REGION Network 249: CARRIER DRIVE INTERNAL COMM ERROR
   RUNG wire#powerrail
      { S7_Templates := "SrcType := Word" } EQ_Contact(in1 := "DB101_DB_SDC_FAULTS".Carrier_Fault[37], in2 := 151)
      Coil( "DB302_HMI_Faults".Carrier37_Faults_1.%X3 )
   END_RUNG
   // the same network as SCL:
   "DB302_HMI_Faults".Carrier37_Faults_1.%X3 := "DB101_DB_SDC_FAULTS".Carrier_Fault[37] = 151;
END_REGION

REGION Network 250: CARRIER DRIVE MOTOR OVERTEMP
   RUNG wire#powerrail
      { S7_Templates := "SrcType := Word" } EQ_Contact(in1 := "DB101_DB_SDC_FAULTS".Carrier_Fault[37], in2 := 160)
      Coil( "DB302_HMI_Faults".Carrier37_Faults_1.%X4 )
   END_RUNG
   // the same network as SCL:
   "DB302_HMI_Faults".Carrier37_Faults_1.%X4 := "DB101_DB_SDC_FAULTS".Carrier_Fault[37] = 160;
END_REGION

REGION Network 251: CARRIER DRIVE MOTOR OVERCURRENT
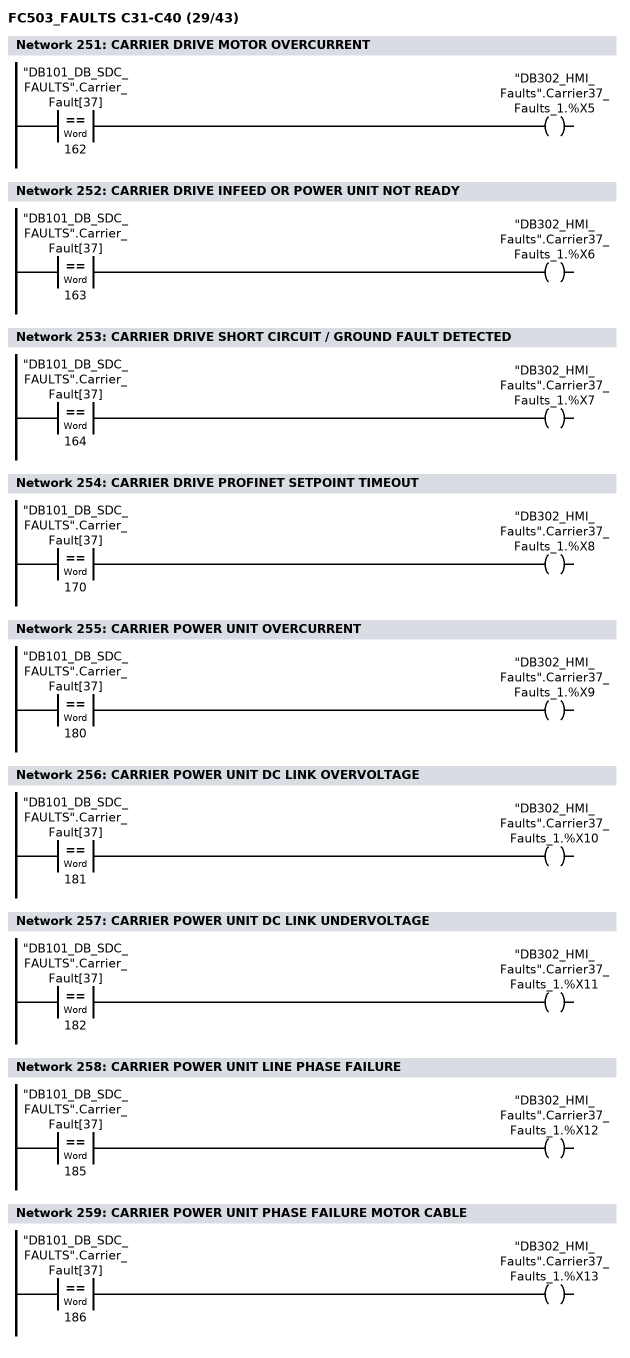
   RUNG wire#powerrail
      { S7_Templates := "SrcType := Word" } EQ_Contact(in1 := "DB101_DB_SDC_FAULTS".Carrier_Fault[37], in2 := 162)
      Coil( "DB302_HMI_Faults".Carrier37_Faults_1.%X5 )
   END_RUNG
   // the same network as SCL:
   "DB302_HMI_Faults".Carrier37_Faults_1.%X5 := "DB101_DB_SDC_FAULTS".Carrier_Fault[37] = 162;
END_REGION

REGION Network 252: CARRIER DRIVE INFEED OR POWER UNIT NOT READY
   RUNG wire#powerrail
      { S7_Templates := "SrcType := Word" } EQ_Contact(in1 := "DB101_DB_SDC_FAULTS".Carrier_Fault[37], in2 := 163)
      Coil( "DB302_HMI_Faults".Carrier37_Faults_1.%X6 )
   END_RUNG
   // the same network as SCL:
   "DB302_HMI_Faults".Carrier37_Faults_1.%X6 := "DB101_DB_SDC_FAULTS".Carrier_Fault[37] = 163;
END_REGION

REGION Network 253: CARRIER DRIVE SHORT CIRCUIT / GROUND FAULT DETECTED
   RUNG wire#powerrail
      { S7_Templates := "SrcType := Word" } EQ_Contact(in1 := "DB101_DB_SDC_FAULTS".Carrier_Fault[37], in2 := 164)
      Coil( "DB302_HMI_Faults".Carrier37_Faults_1.%X7 )
   END_RUNG
   // the same network as SCL:
   "DB302_HMI_Faults".Carrier37_Faults_1.%X7 := "DB101_DB_SDC_FAULTS".Carrier_Fault[37] = 164;
END_REGION

REGION Network 254: CARRIER DRIVE PROFINET SETPOINT TIMEOUT
   RUNG wire#powerrail
      { S7_Templates := "SrcType := Word" } EQ_Contact(in1 := "DB101_DB_SDC_FAULTS".Carrier_Fault[37], in2 := 170)
      Coil( "DB302_HMI_Faults".Carrier37_Faults_1.%X8 )
   END_RUNG
   // the same network as SCL:
   "DB302_HMI_Faults".Carrier37_Faults_1.%X8 := "DB101_DB_SDC_FAULTS".Carrier_Fault[37] = 170;
END_REGION

REGION Network 255: CARRIER POWER UNIT OVERCURRENT
   RUNG wire#powerrail
      { S7_Templates := "SrcType := Word" } EQ_Contact(in1 := "DB101_DB_SDC_FAULTS".Carrier_Fault[37], in2 := 180)
      Coil( "DB302_HMI_Faults".Carrier37_Faults_1.%X9 )
   END_RUNG
   // the same network as SCL:
   "DB302_HMI_Faults".Carrier37_Faults_1.%X9 := "DB101_DB_SDC_FAULTS".Carrier_Fault[37] = 180;
END_REGION

REGION Network 256: CARRIER POWER UNIT DC LINK OVERVOLTAGE
   RUNG wire#powerrail
      { S7_Templates := "SrcType := Word" } EQ_Contact(in1 := "DB101_DB_SDC_FAULTS".Carrier_Fault[37], in2 := 181)
      Coil( "DB302_HMI_Faults".Carrier37_Faults_1.%X10 )
   END_RUNG
   // the same network as SCL:
   "DB302_HMI_Faults".Carrier37_Faults_1.%X10 := "DB101_DB_SDC_FAULTS".Carrier_Fault[37] = 181;
END_REGION

REGION Network 257: CARRIER POWER UNIT DC LINK UNDERVOLTAGE
   RUNG wire#powerrail
      { S7_Templates := "SrcType := Word" } EQ_Contact(in1 := "DB101_DB_SDC_FAULTS".Carrier_Fault[37], in2 := 182)
      Coil( "DB302_HMI_Faults".Carrier37_Faults_1.%X11 )
   END_RUNG
   // the same network as SCL:
   "DB302_HMI_Faults".Carrier37_Faults_1.%X11 := "DB101_DB_SDC_FAULTS".Carrier_Fault[37] = 182;
END_REGION

REGION Network 258: CARRIER POWER UNIT LINE PHASE FAILURE
   RUNG wire#powerrail
      { S7_Templates := "SrcType := Word" } EQ_Contact(in1 := "DB101_DB_SDC_FAULTS".Carrier_Fault[37], in2 := 185)
      Coil( "DB302_HMI_Faults".Carrier37_Faults_1.%X12 )
   END_RUNG
   // the same network as SCL:
   "DB302_HMI_Faults".Carrier37_Faults_1.%X12 := "DB101_DB_SDC_FAULTS".Carrier_Fault[37] = 185;
END_REGION

REGION Network 259: CARRIER POWER UNIT PHASE FAILURE MOTOR CABLE
   RUNG wire#powerrail
      { S7_Templates := "SrcType := Word" } EQ_Contact(in1 := "DB101_DB_SDC_FAULTS".Carrier_Fault[37], in2 := 186)
      Coil( "DB302_HMI_Faults".Carrier37_Faults_1.%X13 )
   END_RUNG
   // the same network as SCL:
   "DB302_HMI_Faults".Carrier37_Faults_1.%X13 := "DB101_DB_SDC_FAULTS".Carrier_Fault[37] = 186;
END_REGION

REGION Network 260: CARRIER POWER UNIT GROUND FAULT
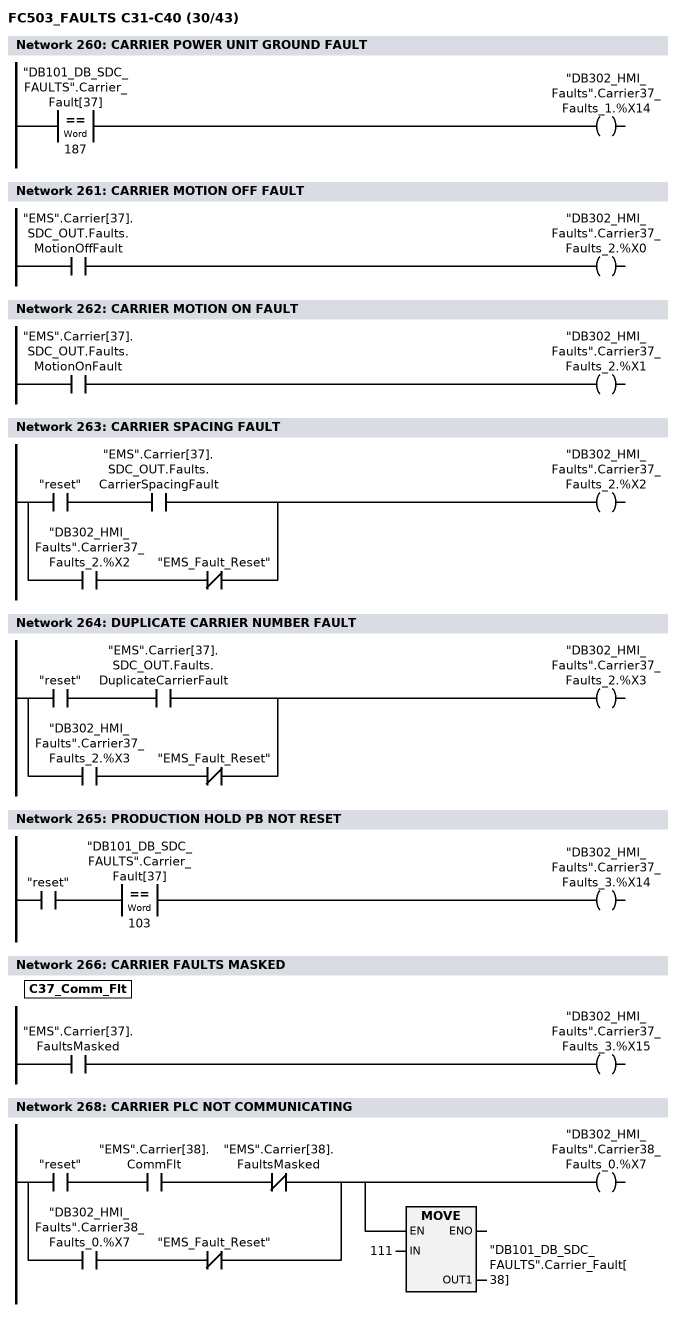
   RUNG wire#powerrail
      { S7_Templates := "SrcType := Word" } EQ_Contact(in1 := "DB101_DB_SDC_FAULTS".Carrier_Fault[37], in2 := 187)
      Coil( "DB302_HMI_Faults".Carrier37_Faults_1.%X14 )
   END_RUNG
   // the same network as SCL:
   "DB302_HMI_Faults".Carrier37_Faults_1.%X14 := "DB101_DB_SDC_FAULTS".Carrier_Fault[37] = 187;
END_REGION

REGION Network 261: CARRIER MOTION OFF FAULT
   RUNG wire#powerrail
      Contact( "EMS".Carrier[37].SDC_OUT.Faults.MotionOffFault )
      Coil( "DB302_HMI_Faults".Carrier37_Faults_2.%X0 )
   END_RUNG
   // the same network as SCL:
   "DB302_HMI_Faults".Carrier37_Faults_2.%X0 := "EMS".Carrier[37].SDC_OUT.Faults.MotionOffFault;
END_REGION

REGION Network 262: CARRIER MOTION ON FAULT
   RUNG wire#powerrail
      Contact( "EMS".Carrier[37].SDC_OUT.Faults.MotionOnFault )
      Coil( "DB302_HMI_Faults".Carrier37_Faults_2.%X1 )
   END_RUNG
   // the same network as SCL:
   "DB302_HMI_Faults".Carrier37_Faults_2.%X1 := "EMS".Carrier[37].SDC_OUT.Faults.MotionOnFault;
END_REGION

REGION Network 263: CARRIER SPACING FAULT
   RUNG wire#powerrail
      Contact( "reset" )
      Contact( "EMS".Carrier[37].SDC_OUT.Faults.CarrierSpacingFault )
      wire#w1
      Coil( "DB302_HMI_Faults".Carrier37_Faults_2.%X2 )
   END_RUNG
   RUNG wire#powerrail
      Contact( "DB302_HMI_Faults".Carrier37_Faults_2.%X2 )
      I_Contact( "EMS_Fault_Reset" )
   END_RUNG wire#w1
   // the same network as SCL:
   "DB302_HMI_Faults".Carrier37_Faults_2.%X2 := ("reset" AND "EMS".Carrier[37].SDC_OUT.Faults.CarrierSpacingFault) OR ("DB302_HMI_Faults".Carrier37_Faults_2.%X2 AND NOT "EMS_Fault_Reset");
END_REGION

REGION Network 264: DUPLICATE CARRIER NUMBER FAULT
   RUNG wire#powerrail
      Contact( "reset" )
      Contact( "EMS".Carrier[37].SDC_OUT.Faults.DuplicateCarrierFault )
      wire#w1
      Coil( "DB302_HMI_Faults".Carrier37_Faults_2.%X3 )
   END_RUNG
   RUNG wire#powerrail
      Contact( "DB302_HMI_Faults".Carrier37_Faults_2.%X3 )
      I_Contact( "EMS_Fault_Reset" )
   END_RUNG wire#w1
   // the same network as SCL:
   "DB302_HMI_Faults".Carrier37_Faults_2.%X3 := ("reset" AND "EMS".Carrier[37].SDC_OUT.Faults.DuplicateCarrierFault) OR ("DB302_HMI_Faults".Carrier37_Faults_2.%X3 AND NOT "EMS_Fault_Reset");
END_REGION

REGION Network 265: PRODUCTION HOLD PB NOT RESET
   RUNG wire#powerrail
      Contact( "reset" )
      { S7_Templates := "SrcType := Word" } EQ_Contact(in1 := "DB101_DB_SDC_FAULTS".Carrier_Fault[37], in2 := 103)
      Coil( "DB302_HMI_Faults".Carrier37_Faults_3.%X14 )
   END_RUNG
   // the same network as SCL:
   "DB302_HMI_Faults".Carrier37_Faults_3.%X14 := "reset" AND ("DB101_DB_SDC_FAULTS".Carrier_Fault[37] = 103);
END_REGION

REGION Network 266: CARRIER FAULTS MASKED
   Label( C37_Comm_Flt )
   RUNG wire#powerrail
      Contact( "EMS".Carrier[37].FaultsMasked )
      Coil( "DB302_HMI_Faults".Carrier37_Faults_3.%X15 )
   END_RUNG
   // the same network as SCL:
   C37_Comm_Flt:
   "DB302_HMI_Faults".Carrier37_Faults_3.%X15 := "EMS".Carrier[37].FaultsMasked;
END_REGION

REGION Network 267: CARRIER 38 FAULTS
END_REGION

REGION Network 268: CARRIER PLC NOT COMMUNICATING
   RUNG wire#powerrail
      Contact( "reset" )
      Contact( "EMS".Carrier[38].CommFlt )
      I_Contact( "EMS".Carrier[38].FaultsMasked )
      wire#w1
      Coil( "DB302_HMI_Faults".Carrier38_Faults_0.%X7 )
   END_RUNG
   RUNG wire#powerrail
      Contact( "DB302_HMI_Faults".Carrier38_Faults_0.%X7 )
      I_Contact( "EMS_Fault_Reset" )
   END_RUNG wire#w1
   RUNG wire#w1
      Move(in := 111, out1 => "DB101_DB_SDC_FAULTS".Carrier_Fault[38])
   END_RUNG
   // the same network as SCL:
   "DB302_HMI_Faults".Carrier38_Faults_0.%X7 := ("reset" AND "EMS".Carrier[38].CommFlt AND NOT "EMS".Carrier[38].FaultsMasked) OR ("DB302_HMI_Faults".Carrier38_Faults_0.%X7 AND NOT "EMS_Fault_Reset");
   IF "DB302_HMI_Faults".Carrier38_Faults_0.%X7 THEN "DB101_DB_SDC_FAULTS".Carrier_Fault[38] := 111; END_IF;
END_REGION

REGION Network 269
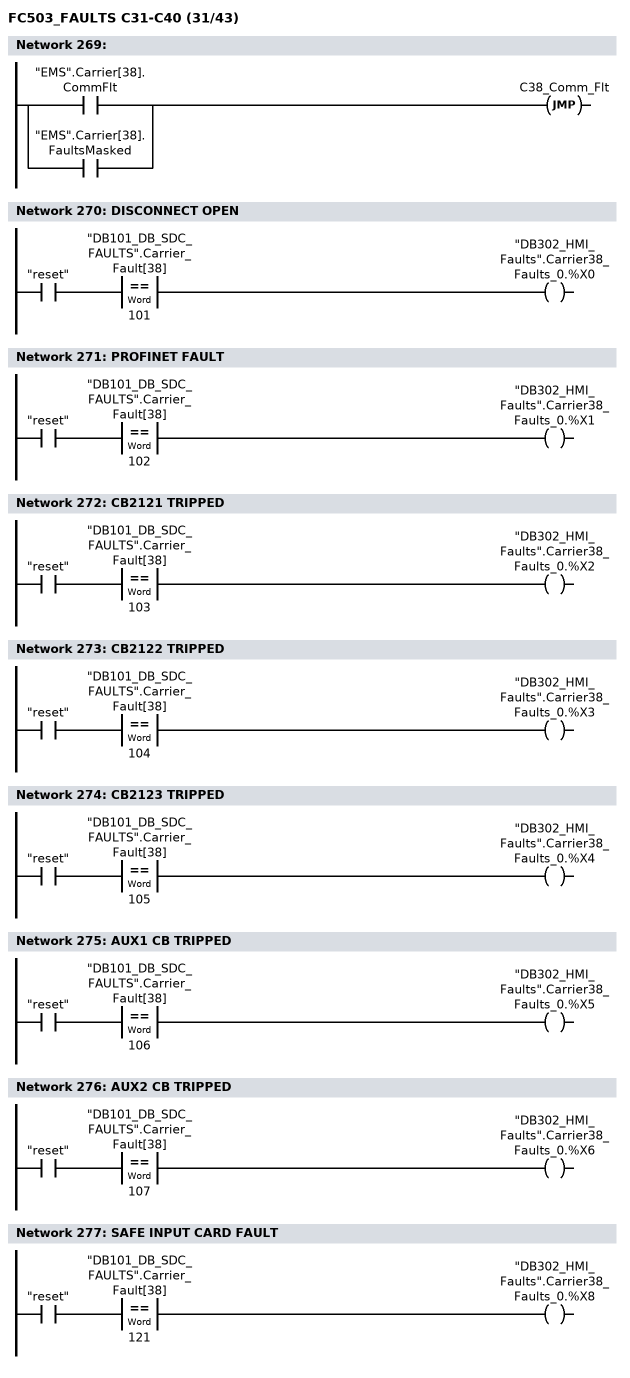
   RUNG wire#powerrail
      Contact( "EMS".Carrier[38].CommFlt )
      wire#w1
      JumpCoil( C38_Comm_Flt )
   END_RUNG
   RUNG wire#powerrail
      Contact( "EMS".Carrier[38].FaultsMasked )
   END_RUNG wire#w1
   // the same network as SCL:
   IF "EMS".Carrier[38].CommFlt OR "EMS".Carrier[38].FaultsMasked THEN GOTO C38_Comm_Flt; END_IF;
END_REGION

REGION Network 270: DISCONNECT OPEN
   RUNG wire#powerrail
      Contact( "reset" )
      { S7_Templates := "SrcType := Word" } EQ_Contact(in1 := "DB101_DB_SDC_FAULTS".Carrier_Fault[38], in2 := 101)
      Coil( "DB302_HMI_Faults".Carrier38_Faults_0.%X0 )
   END_RUNG
   // the same network as SCL:
   "DB302_HMI_Faults".Carrier38_Faults_0.%X0 := "reset" AND ("DB101_DB_SDC_FAULTS".Carrier_Fault[38] = 101);
END_REGION

REGION Network 271: PROFINET FAULT
   RUNG wire#powerrail
      Contact( "reset" )
      { S7_Templates := "SrcType := Word" } EQ_Contact(in1 := "DB101_DB_SDC_FAULTS".Carrier_Fault[38], in2 := 102)
      Coil( "DB302_HMI_Faults".Carrier38_Faults_0.%X1 )
   END_RUNG
   // the same network as SCL:
   "DB302_HMI_Faults".Carrier38_Faults_0.%X1 := "reset" AND ("DB101_DB_SDC_FAULTS".Carrier_Fault[38] = 102);
END_REGION

REGION Network 272: CB2121 TRIPPED
   RUNG wire#powerrail
      Contact( "reset" )
      { S7_Templates := "SrcType := Word" } EQ_Contact(in1 := "DB101_DB_SDC_FAULTS".Carrier_Fault[38], in2 := 103)
      Coil( "DB302_HMI_Faults".Carrier38_Faults_0.%X2 )
   END_RUNG
   // the same network as SCL:
   "DB302_HMI_Faults".Carrier38_Faults_0.%X2 := "reset" AND ("DB101_DB_SDC_FAULTS".Carrier_Fault[38] = 103);
END_REGION

REGION Network 273: CB2122 TRIPPED
   RUNG wire#powerrail
      Contact( "reset" )
      { S7_Templates := "SrcType := Word" } EQ_Contact(in1 := "DB101_DB_SDC_FAULTS".Carrier_Fault[38], in2 := 104)
      Coil( "DB302_HMI_Faults".Carrier38_Faults_0.%X3 )
   END_RUNG
   // the same network as SCL:
   "DB302_HMI_Faults".Carrier38_Faults_0.%X3 := "reset" AND ("DB101_DB_SDC_FAULTS".Carrier_Fault[38] = 104);
END_REGION

REGION Network 274: CB2123 TRIPPED
   RUNG wire#powerrail
      Contact( "reset" )
      { S7_Templates := "SrcType := Word" } EQ_Contact(in1 := "DB101_DB_SDC_FAULTS".Carrier_Fault[38], in2 := 105)
      Coil( "DB302_HMI_Faults".Carrier38_Faults_0.%X4 )
   END_RUNG
   // the same network as SCL:
   "DB302_HMI_Faults".Carrier38_Faults_0.%X4 := "reset" AND ("DB101_DB_SDC_FAULTS".Carrier_Fault[38] = 105);
END_REGION

REGION Network 275: AUX1 CB TRIPPED
   RUNG wire#powerrail
      Contact( "reset" )
      { S7_Templates := "SrcType := Word" } EQ_Contact(in1 := "DB101_DB_SDC_FAULTS".Carrier_Fault[38], in2 := 106)
      Coil( "DB302_HMI_Faults".Carrier38_Faults_0.%X5 )
   END_RUNG
   // the same network as SCL:
   "DB302_HMI_Faults".Carrier38_Faults_0.%X5 := "reset" AND ("DB101_DB_SDC_FAULTS".Carrier_Fault[38] = 106);
END_REGION

REGION Network 276: AUX2 CB TRIPPED
   RUNG wire#powerrail
      Contact( "reset" )
      { S7_Templates := "SrcType := Word" } EQ_Contact(in1 := "DB101_DB_SDC_FAULTS".Carrier_Fault[38], in2 := 107)
      Coil( "DB302_HMI_Faults".Carrier38_Faults_0.%X6 )
   END_RUNG
   // the same network as SCL:
   "DB302_HMI_Faults".Carrier38_Faults_0.%X6 := "reset" AND ("DB101_DB_SDC_FAULTS".Carrier_Fault[38] = 107);
END_REGION

REGION Network 277: SAFE INPUT CARD FAULT
   RUNG wire#powerrail
      Contact( "reset" )
      { S7_Templates := "SrcType := Word" } EQ_Contact(in1 := "DB101_DB_SDC_FAULTS".Carrier_Fault[38], in2 := 121)
      Coil( "DB302_HMI_Faults".Carrier38_Faults_0.%X8 )
   END_RUNG
   // the same network as SCL:
   "DB302_HMI_Faults".Carrier38_Faults_0.%X8 := "reset" AND ("DB101_DB_SDC_FAULTS".Carrier_Fault[38] = 121);
END_REGION

REGION Network 278: SAFE OUTPUT CARD FAULT
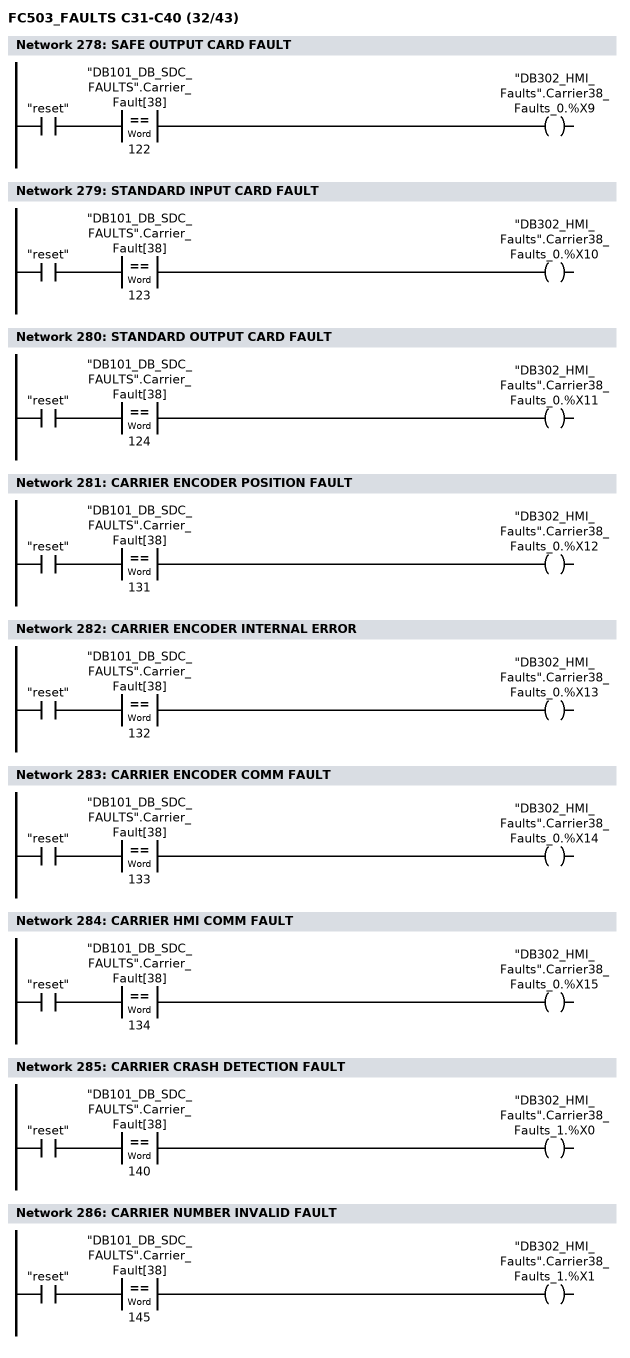
   RUNG wire#powerrail
      Contact( "reset" )
      { S7_Templates := "SrcType := Word" } EQ_Contact(in1 := "DB101_DB_SDC_FAULTS".Carrier_Fault[38], in2 := 122)
      Coil( "DB302_HMI_Faults".Carrier38_Faults_0.%X9 )
   END_RUNG
   // the same network as SCL:
   "DB302_HMI_Faults".Carrier38_Faults_0.%X9 := "reset" AND ("DB101_DB_SDC_FAULTS".Carrier_Fault[38] = 122);
END_REGION

REGION Network 279: STANDARD INPUT CARD FAULT
   RUNG wire#powerrail
      Contact( "reset" )
      { S7_Templates := "SrcType := Word" } EQ_Contact(in1 := "DB101_DB_SDC_FAULTS".Carrier_Fault[38], in2 := 123)
      Coil( "DB302_HMI_Faults".Carrier38_Faults_0.%X10 )
   END_RUNG
   // the same network as SCL:
   "DB302_HMI_Faults".Carrier38_Faults_0.%X10 := "reset" AND ("DB101_DB_SDC_FAULTS".Carrier_Fault[38] = 123);
END_REGION

REGION Network 280: STANDARD OUTPUT CARD FAULT
   RUNG wire#powerrail
      Contact( "reset" )
      { S7_Templates := "SrcType := Word" } EQ_Contact(in1 := "DB101_DB_SDC_FAULTS".Carrier_Fault[38], in2 := 124)
      Coil( "DB302_HMI_Faults".Carrier38_Faults_0.%X11 )
   END_RUNG
   // the same network as SCL:
   "DB302_HMI_Faults".Carrier38_Faults_0.%X11 := "reset" AND ("DB101_DB_SDC_FAULTS".Carrier_Fault[38] = 124);
END_REGION

REGION Network 281: CARRIER ENCODER POSITION FAULT
   RUNG wire#powerrail
      Contact( "reset" )
      { S7_Templates := "SrcType := Word" } EQ_Contact(in1 := "DB101_DB_SDC_FAULTS".Carrier_Fault[38], in2 := 131)
      Coil( "DB302_HMI_Faults".Carrier38_Faults_0.%X12 )
   END_RUNG
   // the same network as SCL:
   "DB302_HMI_Faults".Carrier38_Faults_0.%X12 := "reset" AND ("DB101_DB_SDC_FAULTS".Carrier_Fault[38] = 131);
END_REGION

REGION Network 282: CARRIER ENCODER INTERNAL ERROR
   RUNG wire#powerrail
      Contact( "reset" )
      { S7_Templates := "SrcType := Word" } EQ_Contact(in1 := "DB101_DB_SDC_FAULTS".Carrier_Fault[38], in2 := 132)
      Coil( "DB302_HMI_Faults".Carrier38_Faults_0.%X13 )
   END_RUNG
   // the same network as SCL:
   "DB302_HMI_Faults".Carrier38_Faults_0.%X13 := "reset" AND ("DB101_DB_SDC_FAULTS".Carrier_Fault[38] = 132);
END_REGION

REGION Network 283: CARRIER ENCODER COMM FAULT
   RUNG wire#powerrail
      Contact( "reset" )
      { S7_Templates := "SrcType := Word" } EQ_Contact(in1 := "DB101_DB_SDC_FAULTS".Carrier_Fault[38], in2 := 133)
      Coil( "DB302_HMI_Faults".Carrier38_Faults_0.%X14 )
   END_RUNG
   // the same network as SCL:
   "DB302_HMI_Faults".Carrier38_Faults_0.%X14 := "reset" AND ("DB101_DB_SDC_FAULTS".Carrier_Fault[38] = 133);
END_REGION

REGION Network 284: CARRIER HMI COMM FAULT
   RUNG wire#powerrail
      Contact( "reset" )
      { S7_Templates := "SrcType := Word" } EQ_Contact(in1 := "DB101_DB_SDC_FAULTS".Carrier_Fault[38], in2 := 134)
      Coil( "DB302_HMI_Faults".Carrier38_Faults_0.%X15 )
   END_RUNG
   // the same network as SCL:
   "DB302_HMI_Faults".Carrier38_Faults_0.%X15 := "reset" AND ("DB101_DB_SDC_FAULTS".Carrier_Fault[38] = 134);
END_REGION

REGION Network 285: CARRIER CRASH DETECTION FAULT
   RUNG wire#powerrail
      Contact( "reset" )
      { S7_Templates := "SrcType := Word" } EQ_Contact(in1 := "DB101_DB_SDC_FAULTS".Carrier_Fault[38], in2 := 140)
      Coil( "DB302_HMI_Faults".Carrier38_Faults_1.%X0 )
   END_RUNG
   // the same network as SCL:
   "DB302_HMI_Faults".Carrier38_Faults_1.%X0 := "reset" AND ("DB101_DB_SDC_FAULTS".Carrier_Fault[38] = 140);
END_REGION

REGION Network 286: CARRIER NUMBER INVALID FAULT
   RUNG wire#powerrail
      Contact( "reset" )
      { S7_Templates := "SrcType := Word" } EQ_Contact(in1 := "DB101_DB_SDC_FAULTS".Carrier_Fault[38], in2 := 145)
      Coil( "DB302_HMI_Faults".Carrier38_Faults_1.%X1 )
   END_RUNG
   // the same network as SCL:
   "DB302_HMI_Faults".Carrier38_Faults_1.%X1 := "reset" AND ("DB101_DB_SDC_FAULTS".Carrier_Fault[38] = 145);
END_REGION

REGION Network 287: CARRIER DRIVE PROFINET CONFIG ERROR
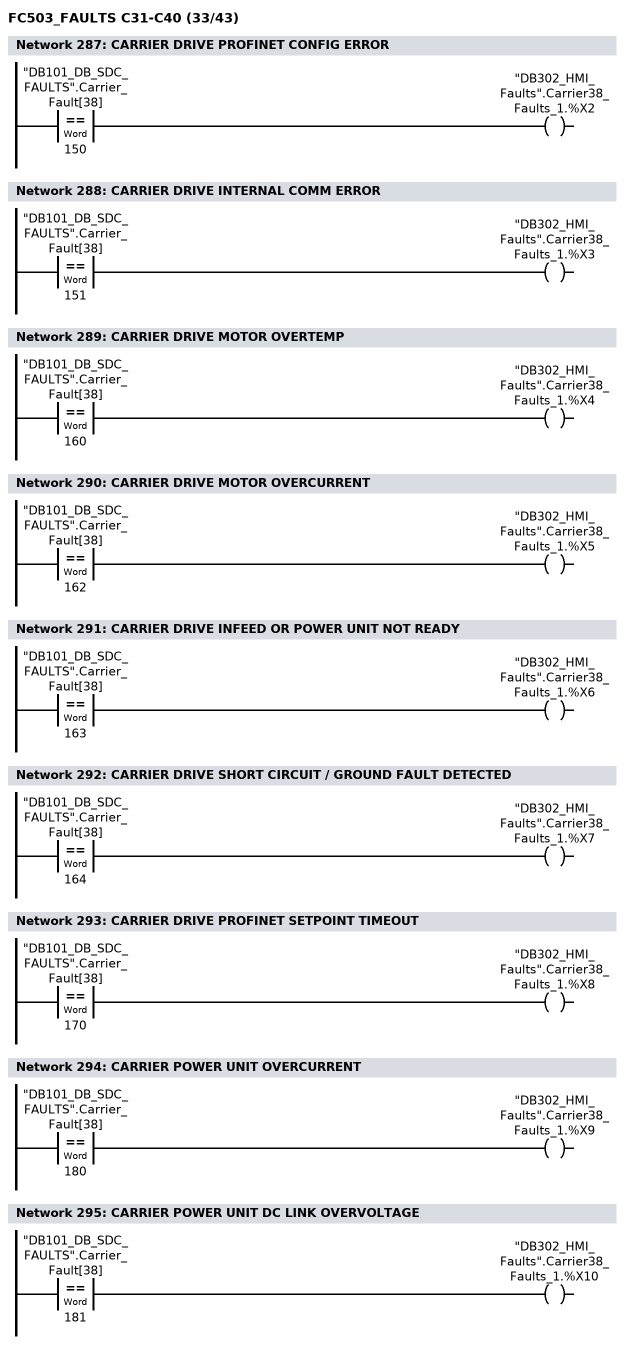
   RUNG wire#powerrail
      { S7_Templates := "SrcType := Word" } EQ_Contact(in1 := "DB101_DB_SDC_FAULTS".Carrier_Fault[38], in2 := 150)
      Coil( "DB302_HMI_Faults".Carrier38_Faults_1.%X2 )
   END_RUNG
   // the same network as SCL:
   "DB302_HMI_Faults".Carrier38_Faults_1.%X2 := "DB101_DB_SDC_FAULTS".Carrier_Fault[38] = 150;
END_REGION

REGION Network 288: CARRIER DRIVE INTERNAL COMM ERROR
   RUNG wire#powerrail
      { S7_Templates := "SrcType := Word" } EQ_Contact(in1 := "DB101_DB_SDC_FAULTS".Carrier_Fault[38], in2 := 151)
      Coil( "DB302_HMI_Faults".Carrier38_Faults_1.%X3 )
   END_RUNG
   // the same network as SCL:
   "DB302_HMI_Faults".Carrier38_Faults_1.%X3 := "DB101_DB_SDC_FAULTS".Carrier_Fault[38] = 151;
END_REGION

REGION Network 289: CARRIER DRIVE MOTOR OVERTEMP
   RUNG wire#powerrail
      { S7_Templates := "SrcType := Word" } EQ_Contact(in1 := "DB101_DB_SDC_FAULTS".Carrier_Fault[38], in2 := 160)
      Coil( "DB302_HMI_Faults".Carrier38_Faults_1.%X4 )
   END_RUNG
   // the same network as SCL:
   "DB302_HMI_Faults".Carrier38_Faults_1.%X4 := "DB101_DB_SDC_FAULTS".Carrier_Fault[38] = 160;
END_REGION

REGION Network 290: CARRIER DRIVE MOTOR OVERCURRENT
   RUNG wire#powerrail
      { S7_Templates := "SrcType := Word" } EQ_Contact(in1 := "DB101_DB_SDC_FAULTS".Carrier_Fault[38], in2 := 162)
      Coil( "DB302_HMI_Faults".Carrier38_Faults_1.%X5 )
   END_RUNG
   // the same network as SCL:
   "DB302_HMI_Faults".Carrier38_Faults_1.%X5 := "DB101_DB_SDC_FAULTS".Carrier_Fault[38] = 162;
END_REGION

REGION Network 291: CARRIER DRIVE INFEED OR POWER UNIT NOT READY
   RUNG wire#powerrail
      { S7_Templates := "SrcType := Word" } EQ_Contact(in1 := "DB101_DB_SDC_FAULTS".Carrier_Fault[38], in2 := 163)
      Coil( "DB302_HMI_Faults".Carrier38_Faults_1.%X6 )
   END_RUNG
   // the same network as SCL:
   "DB302_HMI_Faults".Carrier38_Faults_1.%X6 := "DB101_DB_SDC_FAULTS".Carrier_Fault[38] = 163;
END_REGION

REGION Network 292: CARRIER DRIVE SHORT CIRCUIT / GROUND FAULT DETECTED
   RUNG wire#powerrail
      { S7_Templates := "SrcType := Word" } EQ_Contact(in1 := "DB101_DB_SDC_FAULTS".Carrier_Fault[38], in2 := 164)
      Coil( "DB302_HMI_Faults".Carrier38_Faults_1.%X7 )
   END_RUNG
   // the same network as SCL:
   "DB302_HMI_Faults".Carrier38_Faults_1.%X7 := "DB101_DB_SDC_FAULTS".Carrier_Fault[38] = 164;
END_REGION

REGION Network 293: CARRIER DRIVE PROFINET SETPOINT TIMEOUT
   RUNG wire#powerrail
      { S7_Templates := "SrcType := Word" } EQ_Contact(in1 := "DB101_DB_SDC_FAULTS".Carrier_Fault[38], in2 := 170)
      Coil( "DB302_HMI_Faults".Carrier38_Faults_1.%X8 )
   END_RUNG
   // the same network as SCL:
   "DB302_HMI_Faults".Carrier38_Faults_1.%X8 := "DB101_DB_SDC_FAULTS".Carrier_Fault[38] = 170;
END_REGION

REGION Network 294: CARRIER POWER UNIT OVERCURRENT
   RUNG wire#powerrail
      { S7_Templates := "SrcType := Word" } EQ_Contact(in1 := "DB101_DB_SDC_FAULTS".Carrier_Fault[38], in2 := 180)
      Coil( "DB302_HMI_Faults".Carrier38_Faults_1.%X9 )
   END_RUNG
   // the same network as SCL:
   "DB302_HMI_Faults".Carrier38_Faults_1.%X9 := "DB101_DB_SDC_FAULTS".Carrier_Fault[38] = 180;
END_REGION

REGION Network 295: CARRIER POWER UNIT DC LINK OVERVOLTAGE
   RUNG wire#powerrail
      { S7_Templates := "SrcType := Word" } EQ_Contact(in1 := "DB101_DB_SDC_FAULTS".Carrier_Fault[38], in2 := 181)
      Coil( "DB302_HMI_Faults".Carrier38_Faults_1.%X10 )
   END_RUNG
   // the same network as SCL:
   "DB302_HMI_Faults".Carrier38_Faults_1.%X10 := "DB101_DB_SDC_FAULTS".Carrier_Fault[38] = 181;
END_REGION

REGION Network 296: CARRIER POWER UNIT DC LINK UNDERVOLTAGE
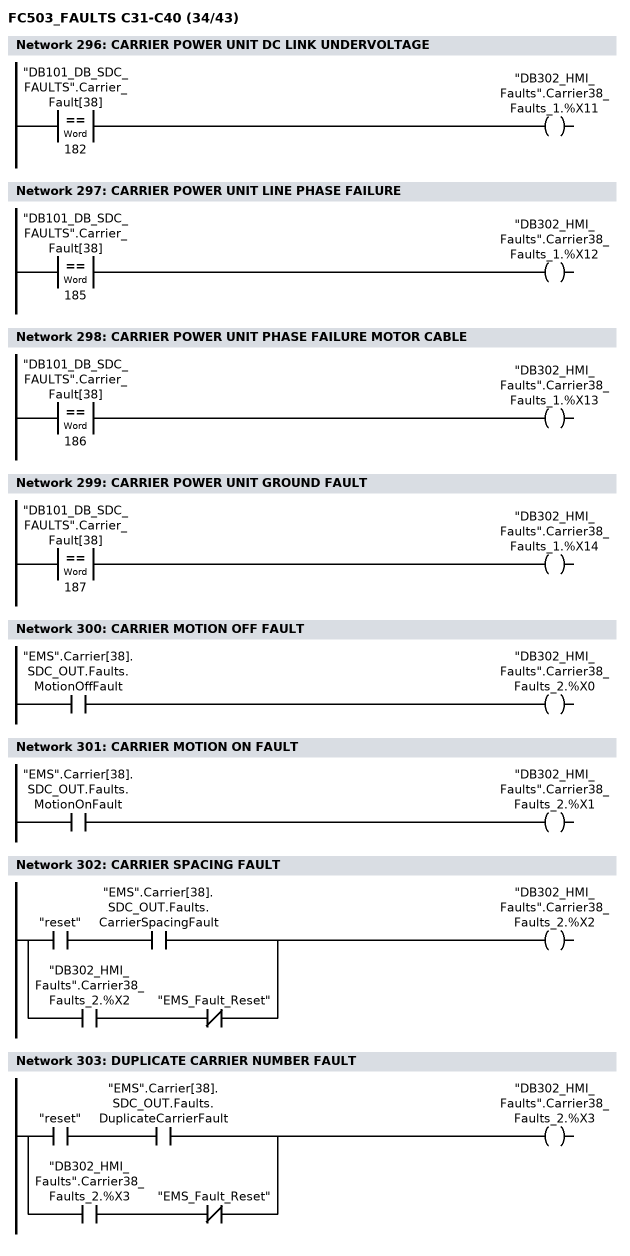
   RUNG wire#powerrail
      { S7_Templates := "SrcType := Word" } EQ_Contact(in1 := "DB101_DB_SDC_FAULTS".Carrier_Fault[38], in2 := 182)
      Coil( "DB302_HMI_Faults".Carrier38_Faults_1.%X11 )
   END_RUNG
   // the same network as SCL:
   "DB302_HMI_Faults".Carrier38_Faults_1.%X11 := "DB101_DB_SDC_FAULTS".Carrier_Fault[38] = 182;
END_REGION

REGION Network 297: CARRIER POWER UNIT LINE PHASE FAILURE
   RUNG wire#powerrail
      { S7_Templates := "SrcType := Word" } EQ_Contact(in1 := "DB101_DB_SDC_FAULTS".Carrier_Fault[38], in2 := 185)
      Coil( "DB302_HMI_Faults".Carrier38_Faults_1.%X12 )
   END_RUNG
   // the same network as SCL:
   "DB302_HMI_Faults".Carrier38_Faults_1.%X12 := "DB101_DB_SDC_FAULTS".Carrier_Fault[38] = 185;
END_REGION

REGION Network 298: CARRIER POWER UNIT PHASE FAILURE MOTOR CABLE
   RUNG wire#powerrail
      { S7_Templates := "SrcType := Word" } EQ_Contact(in1 := "DB101_DB_SDC_FAULTS".Carrier_Fault[38], in2 := 186)
      Coil( "DB302_HMI_Faults".Carrier38_Faults_1.%X13 )
   END_RUNG
   // the same network as SCL:
   "DB302_HMI_Faults".Carrier38_Faults_1.%X13 := "DB101_DB_SDC_FAULTS".Carrier_Fault[38] = 186;
END_REGION

REGION Network 299: CARRIER POWER UNIT GROUND FAULT
   RUNG wire#powerrail
      { S7_Templates := "SrcType := Word" } EQ_Contact(in1 := "DB101_DB_SDC_FAULTS".Carrier_Fault[38], in2 := 187)
      Coil( "DB302_HMI_Faults".Carrier38_Faults_1.%X14 )
   END_RUNG
   // the same network as SCL:
   "DB302_HMI_Faults".Carrier38_Faults_1.%X14 := "DB101_DB_SDC_FAULTS".Carrier_Fault[38] = 187;
END_REGION

REGION Network 300: CARRIER MOTION OFF FAULT
   RUNG wire#powerrail
      Contact( "EMS".Carrier[38].SDC_OUT.Faults.MotionOffFault )
      Coil( "DB302_HMI_Faults".Carrier38_Faults_2.%X0 )
   END_RUNG
   // the same network as SCL:
   "DB302_HMI_Faults".Carrier38_Faults_2.%X0 := "EMS".Carrier[38].SDC_OUT.Faults.MotionOffFault;
END_REGION

REGION Network 301: CARRIER MOTION ON FAULT
   RUNG wire#powerrail
      Contact( "EMS".Carrier[38].SDC_OUT.Faults.MotionOnFault )
      Coil( "DB302_HMI_Faults".Carrier38_Faults_2.%X1 )
   END_RUNG
   // the same network as SCL:
   "DB302_HMI_Faults".Carrier38_Faults_2.%X1 := "EMS".Carrier[38].SDC_OUT.Faults.MotionOnFault;
END_REGION

REGION Network 302: CARRIER SPACING FAULT
   RUNG wire#powerrail
      Contact( "reset" )
      Contact( "EMS".Carrier[38].SDC_OUT.Faults.CarrierSpacingFault )
      wire#w1
      Coil( "DB302_HMI_Faults".Carrier38_Faults_2.%X2 )
   END_RUNG
   RUNG wire#powerrail
      Contact( "DB302_HMI_Faults".Carrier38_Faults_2.%X2 )
      I_Contact( "EMS_Fault_Reset" )
   END_RUNG wire#w1
   // the same network as SCL:
   "DB302_HMI_Faults".Carrier38_Faults_2.%X2 := ("reset" AND "EMS".Carrier[38].SDC_OUT.Faults.CarrierSpacingFault) OR ("DB302_HMI_Faults".Carrier38_Faults_2.%X2 AND NOT "EMS_Fault_Reset");
END_REGION

REGION Network 303: DUPLICATE CARRIER NUMBER FAULT
   RUNG wire#powerrail
      Contact( "reset" )
      Contact( "EMS".Carrier[38].SDC_OUT.Faults.DuplicateCarrierFault )
      wire#w1
      Coil( "DB302_HMI_Faults".Carrier38_Faults_2.%X3 )
   END_RUNG
   RUNG wire#powerrail
      Contact( "DB302_HMI_Faults".Carrier38_Faults_2.%X3 )
      I_Contact( "EMS_Fault_Reset" )
   END_RUNG wire#w1
   // the same network as SCL:
   "DB302_HMI_Faults".Carrier38_Faults_2.%X3 := ("reset" AND "EMS".Carrier[38].SDC_OUT.Faults.DuplicateCarrierFault) OR ("DB302_HMI_Faults".Carrier38_Faults_2.%X3 AND NOT "EMS_Fault_Reset");
END_REGION

REGION Network 304: PRODUCTION HOLD PB NOT RESET
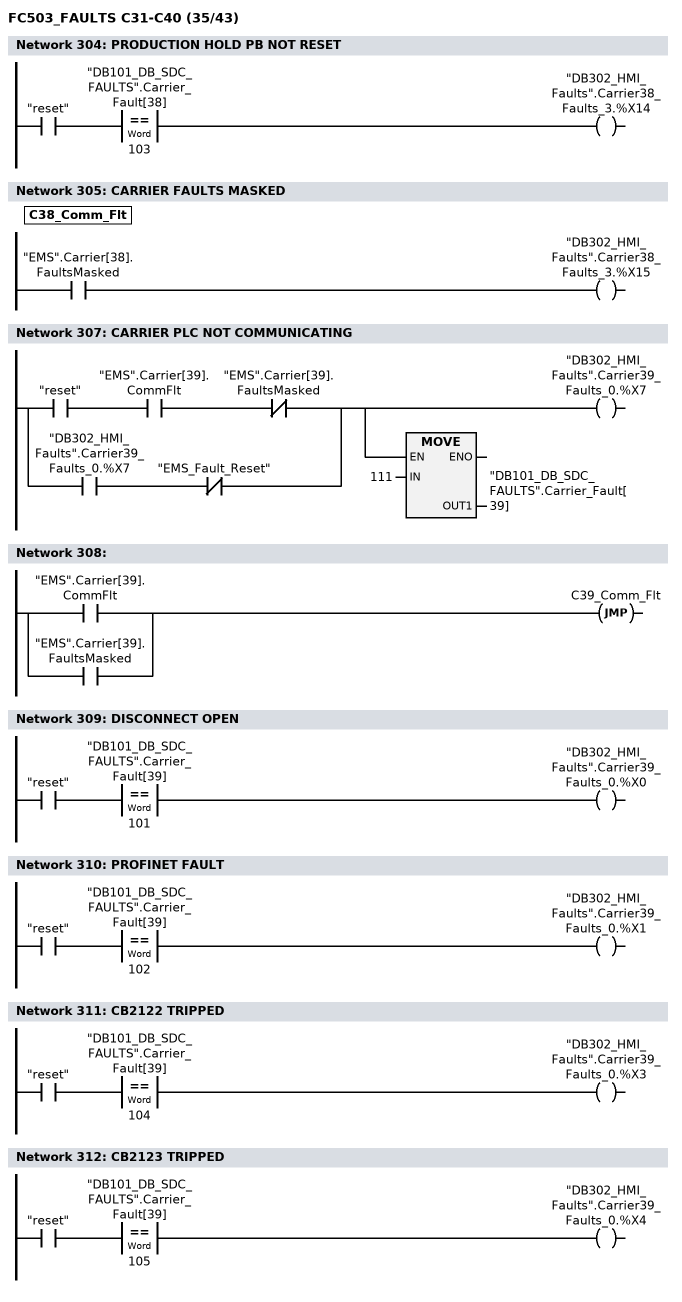
   RUNG wire#powerrail
      Contact( "reset" )
      { S7_Templates := "SrcType := Word" } EQ_Contact(in1 := "DB101_DB_SDC_FAULTS".Carrier_Fault[38], in2 := 103)
      Coil( "DB302_HMI_Faults".Carrier38_Faults_3.%X14 )
   END_RUNG
   // the same network as SCL:
   "DB302_HMI_Faults".Carrier38_Faults_3.%X14 := "reset" AND ("DB101_DB_SDC_FAULTS".Carrier_Fault[38] = 103);
END_REGION

REGION Network 305: CARRIER FAULTS MASKED
   Label( C38_Comm_Flt )
   RUNG wire#powerrail
      Contact( "EMS".Carrier[38].FaultsMasked )
      Coil( "DB302_HMI_Faults".Carrier38_Faults_3.%X15 )
   END_RUNG
   // the same network as SCL:
   C38_Comm_Flt:
   "DB302_HMI_Faults".Carrier38_Faults_3.%X15 := "EMS".Carrier[38].FaultsMasked;
END_REGION

REGION Network 306: CARRIER 39 FAULTS
END_REGION

REGION Network 307: CARRIER PLC NOT COMMUNICATING
   RUNG wire#powerrail
      Contact( "reset" )
      Contact( "EMS".Carrier[39].CommFlt )
      I_Contact( "EMS".Carrier[39].FaultsMasked )
      wire#w1
      Coil( "DB302_HMI_Faults".Carrier39_Faults_0.%X7 )
   END_RUNG
   RUNG wire#powerrail
      Contact( "DB302_HMI_Faults".Carrier39_Faults_0.%X7 )
      I_Contact( "EMS_Fault_Reset" )
   END_RUNG wire#w1
   RUNG wire#w1
      Move(in := 111, out1 => "DB101_DB_SDC_FAULTS".Carrier_Fault[39])
   END_RUNG
   // the same network as SCL:
   "DB302_HMI_Faults".Carrier39_Faults_0.%X7 := ("reset" AND "EMS".Carrier[39].CommFlt AND NOT "EMS".Carrier[39].FaultsMasked) OR ("DB302_HMI_Faults".Carrier39_Faults_0.%X7 AND NOT "EMS_Fault_Reset");
   IF "DB302_HMI_Faults".Carrier39_Faults_0.%X7 THEN "DB101_DB_SDC_FAULTS".Carrier_Fault[39] := 111; END_IF;
END_REGION

REGION Network 308
   RUNG wire#powerrail
      Contact( "EMS".Carrier[39].CommFlt )
      wire#w1
      JumpCoil( C39_Comm_Flt )
   END_RUNG
   RUNG wire#powerrail
      Contact( "EMS".Carrier[39].FaultsMasked )
   END_RUNG wire#w1
   // the same network as SCL:
   IF "EMS".Carrier[39].CommFlt OR "EMS".Carrier[39].FaultsMasked THEN GOTO C39_Comm_Flt; END_IF;
END_REGION

REGION Network 309: DISCONNECT OPEN
   RUNG wire#powerrail
      Contact( "reset" )
      { S7_Templates := "SrcType := Word" } EQ_Contact(in1 := "DB101_DB_SDC_FAULTS".Carrier_Fault[39], in2 := 101)
      Coil( "DB302_HMI_Faults".Carrier39_Faults_0.%X0 )
   END_RUNG
   // the same network as SCL:
   "DB302_HMI_Faults".Carrier39_Faults_0.%X0 := "reset" AND ("DB101_DB_SDC_FAULTS".Carrier_Fault[39] = 101);
END_REGION

REGION Network 310: PROFINET FAULT
   RUNG wire#powerrail
      Contact( "reset" )
      { S7_Templates := "SrcType := Word" } EQ_Contact(in1 := "DB101_DB_SDC_FAULTS".Carrier_Fault[39], in2 := 102)
      Coil( "DB302_HMI_Faults".Carrier39_Faults_0.%X1 )
   END_RUNG
   // the same network as SCL:
   "DB302_HMI_Faults".Carrier39_Faults_0.%X1 := "reset" AND ("DB101_DB_SDC_FAULTS".Carrier_Fault[39] = 102);
END_REGION

REGION Network 311: CB2122 TRIPPED
   RUNG wire#powerrail
      Contact( "reset" )
      { S7_Templates := "SrcType := Word" } EQ_Contact(in1 := "DB101_DB_SDC_FAULTS".Carrier_Fault[39], in2 := 104)
      Coil( "DB302_HMI_Faults".Carrier39_Faults_0.%X3 )
   END_RUNG
   // the same network as SCL:
   "DB302_HMI_Faults".Carrier39_Faults_0.%X3 := "reset" AND ("DB101_DB_SDC_FAULTS".Carrier_Fault[39] = 104);
END_REGION

REGION Network 312: CB2123 TRIPPED
   RUNG wire#powerrail
      Contact( "reset" )
      { S7_Templates := "SrcType := Word" } EQ_Contact(in1 := "DB101_DB_SDC_FAULTS".Carrier_Fault[39], in2 := 105)
      Coil( "DB302_HMI_Faults".Carrier39_Faults_0.%X4 )
   END_RUNG
   // the same network as SCL:
   "DB302_HMI_Faults".Carrier39_Faults_0.%X4 := "reset" AND ("DB101_DB_SDC_FAULTS".Carrier_Fault[39] = 105);
END_REGION

REGION Network 313: AUX1 CB TRIPPED
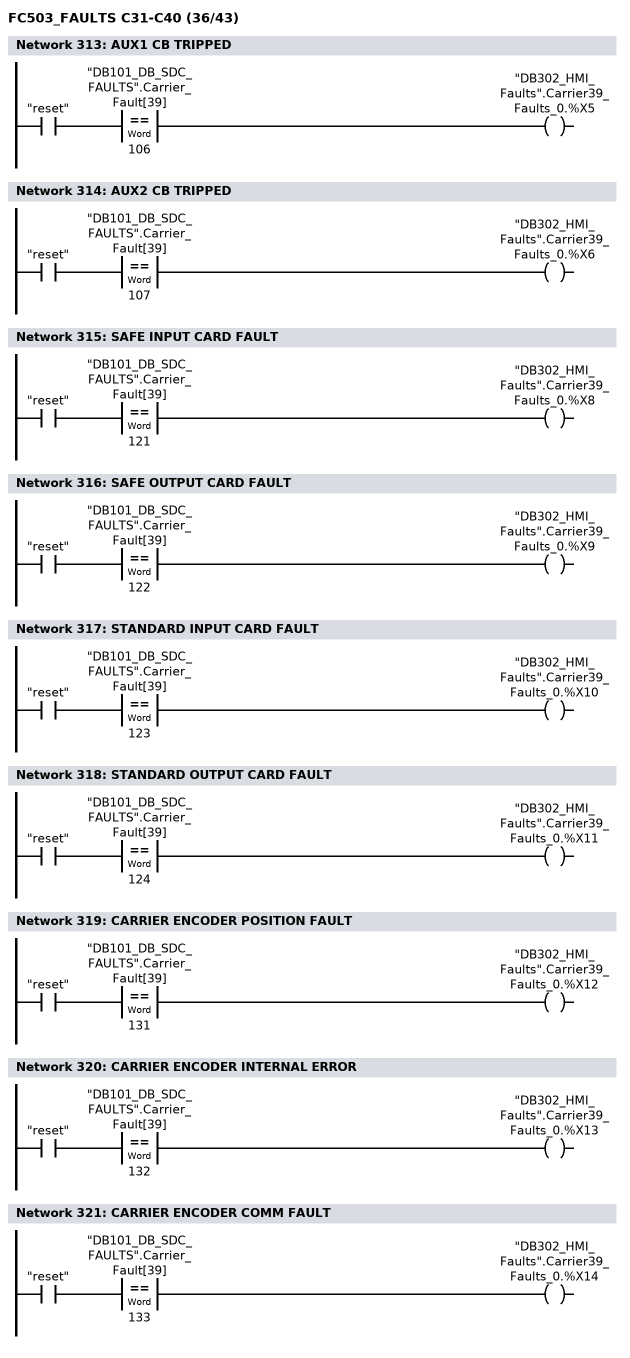
   RUNG wire#powerrail
      Contact( "reset" )
      { S7_Templates := "SrcType := Word" } EQ_Contact(in1 := "DB101_DB_SDC_FAULTS".Carrier_Fault[39], in2 := 106)
      Coil( "DB302_HMI_Faults".Carrier39_Faults_0.%X5 )
   END_RUNG
   // the same network as SCL:
   "DB302_HMI_Faults".Carrier39_Faults_0.%X5 := "reset" AND ("DB101_DB_SDC_FAULTS".Carrier_Fault[39] = 106);
END_REGION

REGION Network 314: AUX2 CB TRIPPED
   RUNG wire#powerrail
      Contact( "reset" )
      { S7_Templates := "SrcType := Word" } EQ_Contact(in1 := "DB101_DB_SDC_FAULTS".Carrier_Fault[39], in2 := 107)
      Coil( "DB302_HMI_Faults".Carrier39_Faults_0.%X6 )
   END_RUNG
   // the same network as SCL:
   "DB302_HMI_Faults".Carrier39_Faults_0.%X6 := "reset" AND ("DB101_DB_SDC_FAULTS".Carrier_Fault[39] = 107);
END_REGION

REGION Network 315: SAFE INPUT CARD FAULT
   RUNG wire#powerrail
      Contact( "reset" )
      { S7_Templates := "SrcType := Word" } EQ_Contact(in1 := "DB101_DB_SDC_FAULTS".Carrier_Fault[39], in2 := 121)
      Coil( "DB302_HMI_Faults".Carrier39_Faults_0.%X8 )
   END_RUNG
   // the same network as SCL:
   "DB302_HMI_Faults".Carrier39_Faults_0.%X8 := "reset" AND ("DB101_DB_SDC_FAULTS".Carrier_Fault[39] = 121);
END_REGION

REGION Network 316: SAFE OUTPUT CARD FAULT
   RUNG wire#powerrail
      Contact( "reset" )
      { S7_Templates := "SrcType := Word" } EQ_Contact(in1 := "DB101_DB_SDC_FAULTS".Carrier_Fault[39], in2 := 122)
      Coil( "DB302_HMI_Faults".Carrier39_Faults_0.%X9 )
   END_RUNG
   // the same network as SCL:
   "DB302_HMI_Faults".Carrier39_Faults_0.%X9 := "reset" AND ("DB101_DB_SDC_FAULTS".Carrier_Fault[39] = 122);
END_REGION

REGION Network 317: STANDARD INPUT CARD FAULT
   RUNG wire#powerrail
      Contact( "reset" )
      { S7_Templates := "SrcType := Word" } EQ_Contact(in1 := "DB101_DB_SDC_FAULTS".Carrier_Fault[39], in2 := 123)
      Coil( "DB302_HMI_Faults".Carrier39_Faults_0.%X10 )
   END_RUNG
   // the same network as SCL:
   "DB302_HMI_Faults".Carrier39_Faults_0.%X10 := "reset" AND ("DB101_DB_SDC_FAULTS".Carrier_Fault[39] = 123);
END_REGION

REGION Network 318: STANDARD OUTPUT CARD FAULT
   RUNG wire#powerrail
      Contact( "reset" )
      { S7_Templates := "SrcType := Word" } EQ_Contact(in1 := "DB101_DB_SDC_FAULTS".Carrier_Fault[39], in2 := 124)
      Coil( "DB302_HMI_Faults".Carrier39_Faults_0.%X11 )
   END_RUNG
   // the same network as SCL:
   "DB302_HMI_Faults".Carrier39_Faults_0.%X11 := "reset" AND ("DB101_DB_SDC_FAULTS".Carrier_Fault[39] = 124);
END_REGION
